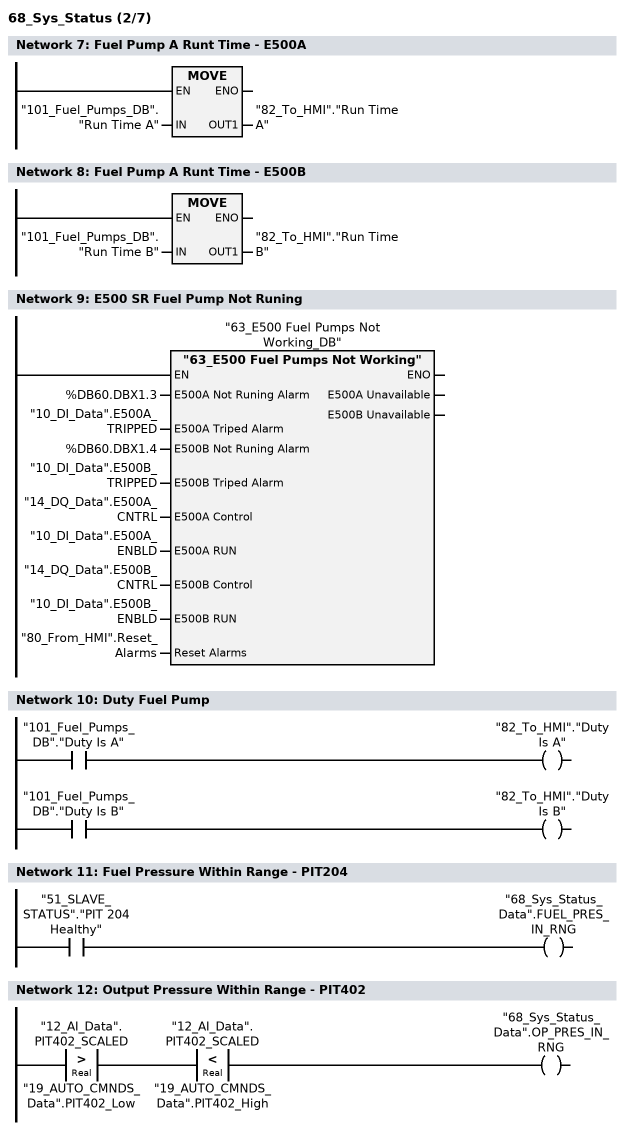
   RUNG wire#powerrail
      Move(in := "101_Fuel_Pumps_DB"."Run Time A", out1 => "82_To_HMI"."Run Time A")
   END_RUNG
   // the same network as SCL:
   "82_To_HMI"."Run Time A" := "101_Fuel_Pumps_DB"."Run Time A";
END_REGION

REGION Network 8: Fuel Pump A Runt Time - E500B
   RUNG wire#powerrail
      Move(in := "101_Fuel_Pumps_DB"."Run Time B", out1 => "82_To_HMI"."Run Time B")
   END_RUNG
   // the same network as SCL:
   "82_To_HMI"."Run Time B" := "101_Fuel_Pumps_DB"."Run Time B";
END_REGION

REGION Network 9: E500 SR Fuel Pump Not Runing
   RUNG wire#powerrail
      "63_E500 Fuel Pumps Not Working_DB"("E500A Not Runing Alarm" := %DB60.DBX1.3, "E500A Triped Alarm" := "10_DI_Data".E500A_TRIPPED, "E500B Not Runing Alarm" := %DB60.DBX1.4, "E500B Triped Alarm" := "10_DI_Data".E500B_TRIPPED, "E500A Control" := "14_DQ_Data".E500A_CNTRL, "E500A RUN" := "10_DI_Data".E500A_ENBLD, "E500B Control" := "14_DQ_Data".E500B_CNTRL, "E500B RUN" := "10_DI_Data".E500B_ENBLD, "Reset Alarms" := "80_From_HMI".Reset_Alarms, "E500A Unavailable" =>, "E500B Unavailable" =>)
   END_RUNG
   // the same network as SCL:
   "63_E500 Fuel Pumps Not Working_DB"("E500A Not Runing Alarm" := %DB60.DBX1.3,   // "63_E500 Fuel Pumps Not Working"
                           "E500A Triped Alarm" := "10_DI_Data".E500A_TRIPPED,
                           "E500B Not Runing Alarm" := %DB60.DBX1.4,
                           "E500B Triped Alarm" := "10_DI_Data".E500B_TRIPPED,
                           "E500A Control" := "14_DQ_Data".E500A_CNTRL,
                           "E500A RUN" := "10_DI_Data".E500A_ENBLD,
                           "E500B Control" := "14_DQ_Data".E500B_CNTRL,
                           "E500B RUN" := "10_DI_Data".E500B_ENBLD,
                           "Reset Alarms" := "80_From_HMI".Reset_Alarms);
END_REGION

REGION Network 10: Duty Fuel Pump
   RUNG wire#powerrail
      Contact( "101_Fuel_Pumps_DB"."Duty Is A" )
      Coil( "82_To_HMI"."Duty Is A" )
   END_RUNG
   RUNG wire#powerrail
      Contact( "101_Fuel_Pumps_DB"."Duty Is B" )
      Coil( "82_To_HMI"."Duty Is B" )
   END_RUNG
   // the same network as SCL:
   "82_To_HMI"."Duty Is A" := "101_Fuel_Pumps_DB"."Duty Is A";
   "82_To_HMI"."Duty Is B" := "101_Fuel_Pumps_DB"."Duty Is B";
END_REGION

REGION Network 11: Fuel Pressure Within Range - PIT204
   RUNG wire#powerrail
      Contact( "51_SLAVE_STATUS"."PIT 204 Healthy" )
      Coil( "68_Sys_Status_Data".FUEL_PRES_IN_RNG )
   END_RUNG
   // the same network as SCL:
   "68_Sys_Status_Data".FUEL_PRES_IN_RNG := "51_SLAVE_STATUS"."PIT 204 Healthy";
END_REGION

REGION Network 12: Output Pressure Within Range - PIT402
   RUNG wire#powerrail
      { S7_Templates := "SrcType := Real" } GT_Contact(in1 := "12_AI_Data".PIT402_SCALED, in2 := "19_AUTO_CMNDS_Data".PIT402_Low)
      { S7_Templates := "SrcType := Real" } LT_Contact(in1 := "12_AI_Data".PIT402_SCALED, in2 := "19_AUTO_CMNDS_Data".PIT402_High)
      Coil( "68_Sys_Status_Data".OP_PRES_IN_RNG )
   END_RUNG
   // the same network as SCL:
   "68_Sys_Status_Data".OP_PRES_IN_RNG := ("12_AI_Data".PIT402_SCALED > "19_AUTO_CMNDS_Data".PIT402_Low) AND ("12_AI_Data".PIT402_SCALED < "19_AUTO_CMNDS_Data".PIT402_High);
END_REGION

REGION Network 13: Cargo Banketing Mode
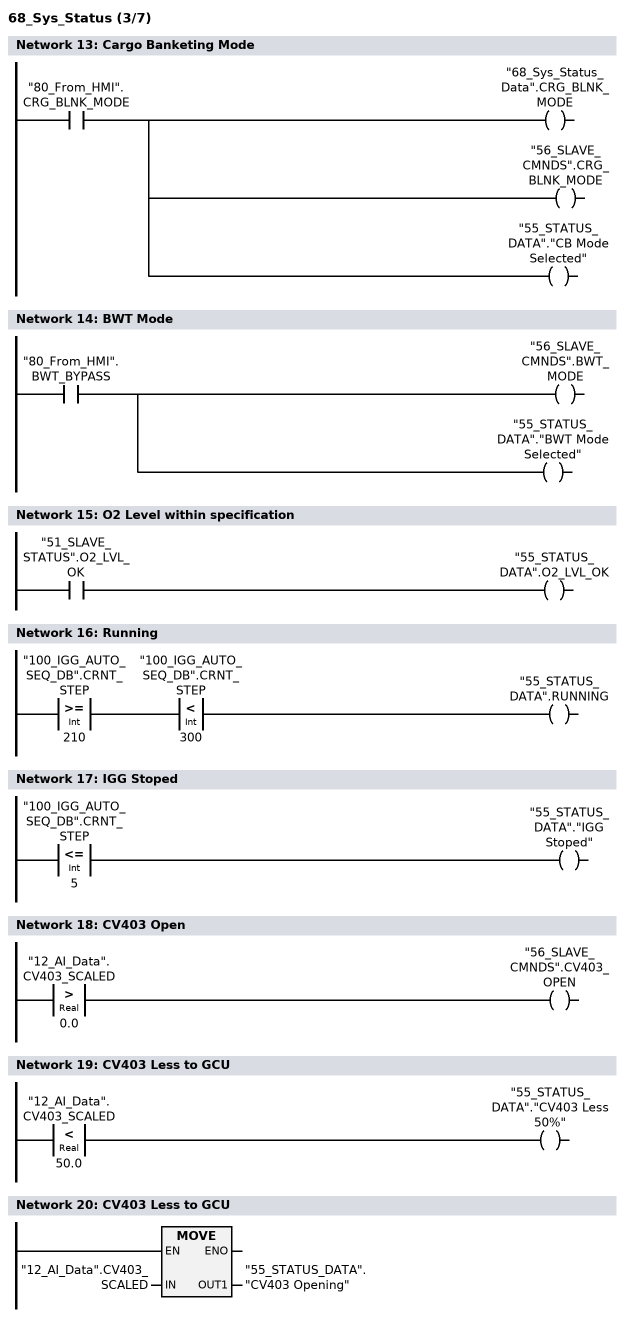
   RUNG wire#powerrail
      Contact( "80_From_HMI".CRG_BLNK_MODE )
      wire#w1
      Coil( "68_Sys_Status_Data".CRG_BLNK_MODE )
   END_RUNG
   RUNG wire#w1
      Coil( "56_SLAVE_CMNDS".CRG_BLNK_MODE )
   END_RUNG
   RUNG wire#w1
      Coil( "55_STATUS_DATA"."CB Mode Selected" )
   END_RUNG
   // the same network as SCL:
   "68_Sys_Status_Data".CRG_BLNK_MODE := "80_From_HMI".CRG_BLNK_MODE;
   "56_SLAVE_CMNDS".CRG_BLNK_MODE := "80_From_HMI".CRG_BLNK_MODE;
   "55_STATUS_DATA"."CB Mode Selected" := "80_From_HMI".CRG_BLNK_MODE;
END_REGION

REGION Network 14: BWT Mode
   RUNG wire#powerrail
      Contact( "80_From_HMI".BWT_BYPASS )
      wire#w1
      Coil( "56_SLAVE_CMNDS".BWT_MODE )
   END_RUNG
   RUNG wire#w1
      Coil( "55_STATUS_DATA"."BWT Mode Selected" )
   END_RUNG
   // the same network as SCL:
   "56_SLAVE_CMNDS".BWT_MODE := "80_From_HMI".BWT_BYPASS;
   "55_STATUS_DATA"."BWT Mode Selected" := "80_From_HMI".BWT_BYPASS;
END_REGION

REGION Network 15: O2 Level within specification
   RUNG wire#powerrail
      Contact( "51_SLAVE_STATUS".O2_LVL_OK )
      Coil( "55_STATUS_DATA".O2_LVL_OK )
   END_RUNG
   // the same network as SCL:
   "55_STATUS_DATA".O2_LVL_OK := "51_SLAVE_STATUS".O2_LVL_OK;
END_REGION

REGION Network 16: Running
   RUNG wire#powerrail
      { S7_Templates := "SrcType := Int" } GE_Contact(in1 := "100_IGG_AUTO_SEQ_DB".CRNT_STEP, in2 := 210)
      { S7_Templates := "SrcType := Int" } LT_Contact(in1 := "100_IGG_AUTO_SEQ_DB".CRNT_STEP, in2 := 300)
      Coil( "55_STATUS_DATA".RUNNING )
   END_RUNG
   // the same network as SCL:
   "55_STATUS_DATA".RUNNING := ("100_IGG_AUTO_SEQ_DB".CRNT_STEP >= 210) AND ("100_IGG_AUTO_SEQ_DB".CRNT_STEP < 300);
END_REGION

REGION Network 17: IGG Stoped
   RUNG wire#powerrail
      { S7_Templates := "SrcType := Int" } LE_Contact(in1 := "100_IGG_AUTO_SEQ_DB".CRNT_STEP, in2 := 5)
      Coil( "55_STATUS_DATA"."IGG Stoped" )
   END_RUNG
   // the same network as SCL:
   "55_STATUS_DATA"."IGG Stoped" := "100_IGG_AUTO_SEQ_DB".CRNT_STEP <= 5;
END_REGION

REGION Network 18: CV403 Open
   RUNG wire#powerrail
      { S7_Templates := "SrcType := Real" } GT_Contact(in1 := "12_AI_Data".CV403_SCALED, in2 := 0.0)
      Coil( "56_SLAVE_CMNDS".CV403_OPEN )
   END_RUNG
   // the same network as SCL:
   "56_SLAVE_CMNDS".CV403_OPEN := "12_AI_Data".CV403_SCALED > 0.0;
END_REGION

REGION Network 19: CV403 Less to GCU
   RUNG wire#powerrail
      { S7_Templates := "SrcType := Real" } LT_Contact(in1 := "12_AI_Data".CV403_SCALED, in2 := 50.0)
      Coil( "55_STATUS_DATA"."CV403 Less 50%" )
   END_RUNG
   // the same network as SCL:
   "55_STATUS_DATA"."CV403 Less 50%" := "12_AI_Data".CV403_SCALED < 50.0;
END_REGION

REGION Network 20: CV403 Less to GCU
   RUNG wire#powerrail
      Move(in := "12_AI_Data".CV403_SCALED, out1 => "55_STATUS_DATA"."CV403 Opening")
   END_RUNG
   // the same network as SCL:
   "55_STATUS_DATA"."CV403 Opening" := "12_AI_Data".CV403_SCALED;
END_REGION

REGION Network 21: Fuel Pump 1 Enabled E500A
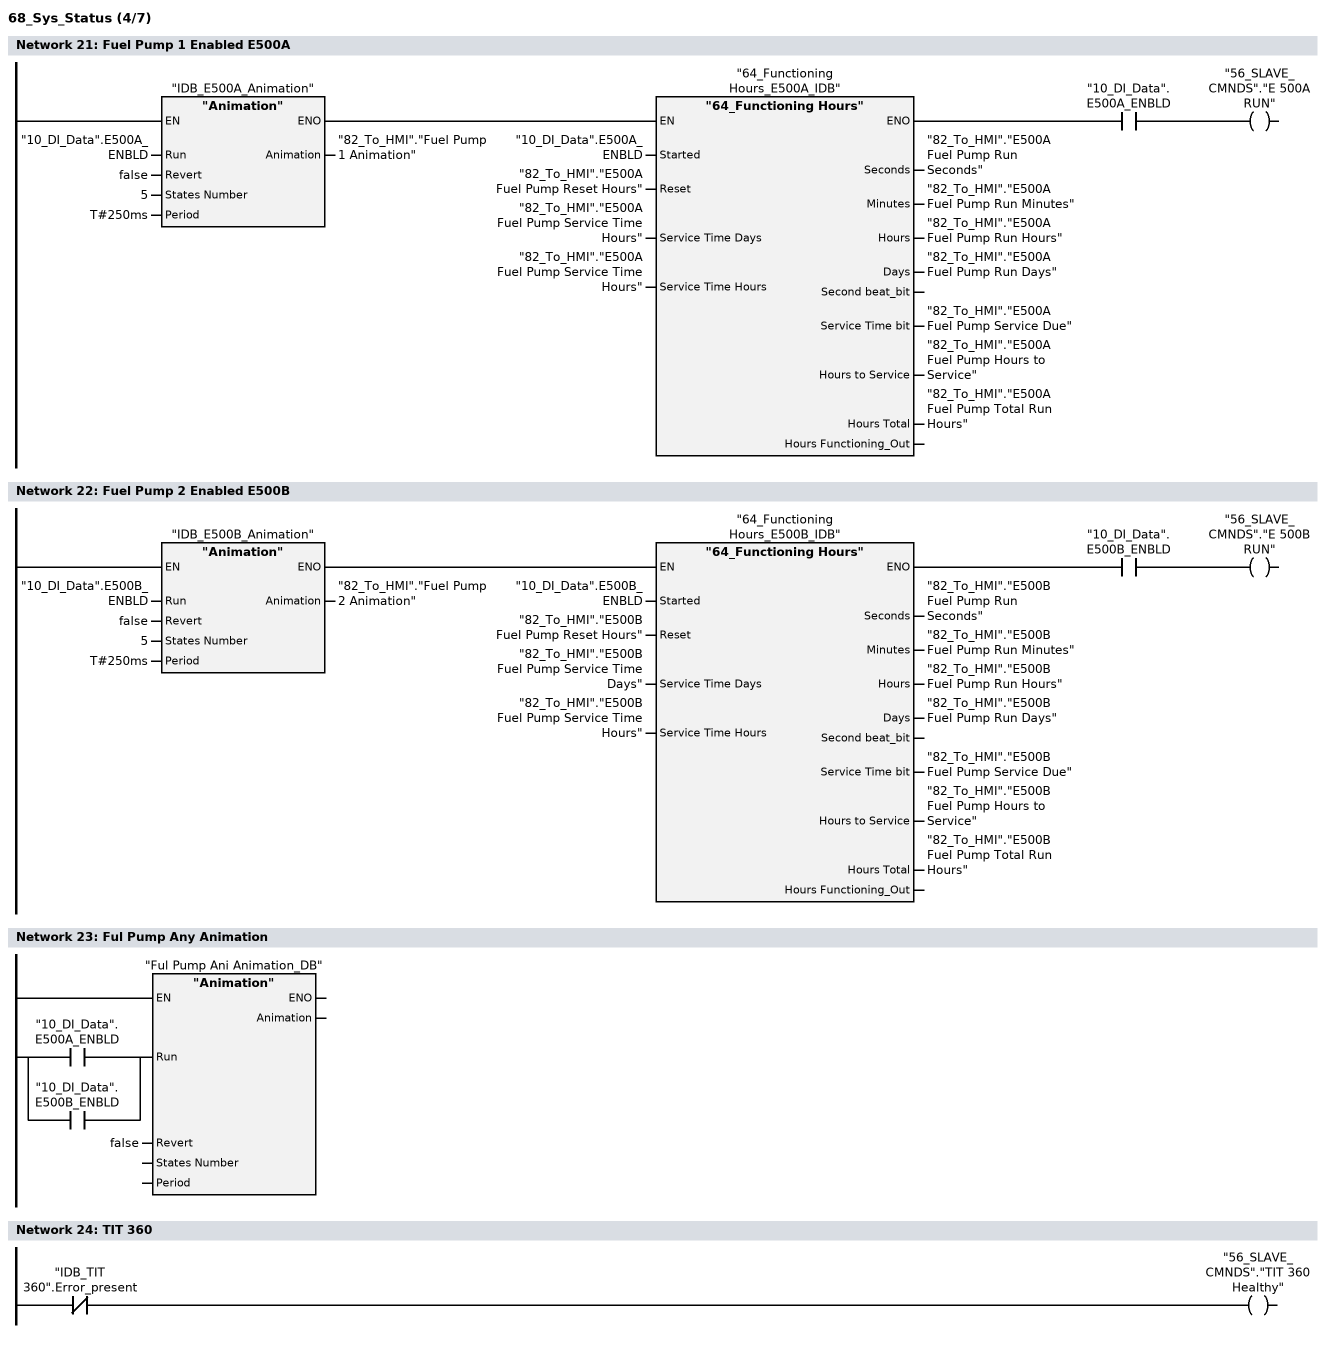
   RUNG wire#powerrail
      "IDB_E500A_Animation"(Run := "10_DI_Data".E500A_ENBLD, Revert := false, "States Number" := 5, Period := T#250ms, Animation => "82_To_HMI"."Fuel Pump 1 Animation")
      "64_Functioning Hours_E500A_IDB"(Started := "10_DI_Data".E500A_ENBLD, Reset := "82_To_HMI"."E500A Fuel Pump Reset Hours", "Service Time Days" := "82_To_HMI"."E500A Fuel Pump Service Time Hours", "Service Time Hours" := "82_To_HMI"."E500A Fuel Pump Service Time Hours", Seconds => "82_To_HMI"."E500A Fuel Pump Run Seconds", Minutes => "82_To_HMI"."E500A Fuel Pump Run Minutes", Hours => "82_To_HMI"."E500A Fuel Pump Run Hours", Days => "82_To_HMI"."E500A Fuel Pump Run Days", "Second beat_bit" =>, "Service Time bit" => "82_To_HMI"."E500A Fuel Pump Service Due", "Hours to Service" => "82_To_HMI"."E500A Fuel Pump Hours to Service", "Hours Total" => "82_To_HMI"."E500A Fuel Pump Total Run Hours", "Hours Functioning_Out" =>)
      Contact( "10_DI_Data".E500A_ENBLD )
      Coil( "56_SLAVE_CMNDS"."E 500A RUN" )
   END_RUNG
   // the same network as SCL:
   "IDB_E500A_Animation"(Run := "10_DI_Data".E500A_ENBLD,   // "Animation"
                         Revert := false,
                         "States Number" := 5,
                         Period := T#250ms,
                         Animation => "82_To_HMI"."Fuel Pump 1 Animation",
                         ENO => #_w1);
   "64_Functioning Hours_E500A_IDB"(EN := #_w1,   // "64_Functioning Hours"
                           Started := "10_DI_Data".E500A_ENBLD,
                           Reset := "82_To_HMI"."E500A Fuel Pump Reset Hours",
                           "Service Time Days" := "82_To_HMI"."E500A Fuel Pump Service Time Hours",
                           "Service Time Hours" := "82_To_HMI"."E500A Fuel Pump Service Time Hours",
                           Seconds => "82_To_HMI"."E500A Fuel Pump Run Seconds",
                           Minutes => "82_To_HMI"."E500A Fuel Pump Run Minutes",
                           Hours => "82_To_HMI"."E500A Fuel Pump Run Hours",
                           Days => "82_To_HMI"."E500A Fuel Pump Run Days",
                           "Service Time bit" => "82_To_HMI"."E500A Fuel Pump Service Due",
                           "Hours to Service" => "82_To_HMI"."E500A Fuel Pump Hours to Service",
                           "Hours Total" => "82_To_HMI"."E500A Fuel Pump Total Run Hours",
                           ENO => #_w2);
   "56_SLAVE_CMNDS"."E 500A RUN" := #_w2 AND "10_DI_Data".E500A_ENBLD;
END_REGION

REGION Network 22: Fuel Pump 2 Enabled E500B
   RUNG wire#powerrail
      "IDB_E500B_Animation"(Run := "10_DI_Data".E500B_ENBLD, Revert := false, "States Number" := 5, Period := T#250ms, Animation => "82_To_HMI"."Fuel Pump 2 Animation")
      "64_Functioning Hours_E500B_IDB"(Started := "10_DI_Data".E500B_ENBLD, Reset := "82_To_HMI"."E500B Fuel Pump Reset Hours", "Service Time Days" := "82_To_HMI"."E500B Fuel Pump Service Time Days", "Service Time Hours" := "82_To_HMI"."E500B Fuel Pump Service Time Hours", Seconds => "82_To_HMI"."E500B Fuel Pump Run Seconds", Minutes => "82_To_HMI"."E500B Fuel Pump Run Minutes", Hours => "82_To_HMI"."E500B Fuel Pump Run Hours", Days => "82_To_HMI"."E500B Fuel Pump Run Days", "Second beat_bit" =>, "Service Time bit" => "82_To_HMI"."E500B Fuel Pump Service Due", "Hours to Service" => "82_To_HMI"."E500B Fuel Pump Hours to Service", "Hours Total" => "82_To_HMI"."E500B Fuel Pump Total Run Hours", "Hours Functioning_Out" =>)
      Contact( "10_DI_Data".E500B_ENBLD )
      Coil( "56_SLAVE_CMNDS"."E 500B RUN" )
   END_RUNG
   // the same network as SCL:
   "IDB_E500B_Animation"(Run := "10_DI_Data".E500B_ENBLD,   // "Animation"
                         Revert := false,
                         "States Number" := 5,
                         Period := T#250ms,
                         Animation => "82_To_HMI"."Fuel Pump 2 Animation",
                         ENO => #_w1);
   "64_Functioning Hours_E500B_IDB"(EN := #_w1,   // "64_Functioning Hours"
                           Started := "10_DI_Data".E500B_ENBLD,
                           Reset := "82_To_HMI"."E500B Fuel Pump Reset Hours",
                           "Service Time Days" := "82_To_HMI"."E500B Fuel Pump Service Time Days",
                           "Service Time Hours" := "82_To_HMI"."E500B Fuel Pump Service Time Hours",
                           Seconds => "82_To_HMI"."E500B Fuel Pump Run Seconds",
                           Minutes => "82_To_HMI"."E500B Fuel Pump Run Minutes",
                           Hours => "82_To_HMI"."E500B Fuel Pump Run Hours",
                           Days => "82_To_HMI"."E500B Fuel Pump Run Days",
                           "Service Time bit" => "82_To_HMI"."E500B Fuel Pump Service Due",
                           "Hours to Service" => "82_To_HMI"."E500B Fuel Pump Hours to Service",
                           "Hours Total" => "82_To_HMI"."E500B Fuel Pump Total Run Hours",
                           ENO => #_w2);
   "56_SLAVE_CMNDS"."E 500B RUN" := #_w2 AND "10_DI_Data".E500B_ENBLD;
END_REGION

REGION Network 23: Ful Pump Any Animation
   RUNG wire#powerrail
      "Ful Pump Ani Animation_DB"(Run := wire#w1, Revert := false, "States Number" :=, Period :=, Animation =>)
   END_RUNG
   RUNG wire#powerrail
      Contact( "10_DI_Data".E500A_ENBLD )
   END_RUNG wire#w1
   RUNG wire#powerrail
      Contact( "10_DI_Data".E500B_ENBLD )
   END_RUNG wire#w1
   // the same network as SCL:
   "Ful Pump Ani Animation_DB"(Run := "10_DI_Data".E500A_ENBLD OR "10_DI_Data".E500B_ENBLD, Revert := false);   // "Animation"
END_REGION

REGION Network 24: TIT 360
   RUNG wire#powerrail
      I_Contact( "IDB_TIT 360".Error_present )
      Coil( "56_SLAVE_CMNDS"."TIT 360 Healthy" )
   END_RUNG
   // the same network as SCL:
   "56_SLAVE_CMNDS"."TIT 360 Healthy" := NOT "IDB_TIT 360".Error_present;
END_REGION

REGION Network 25: TIT 401
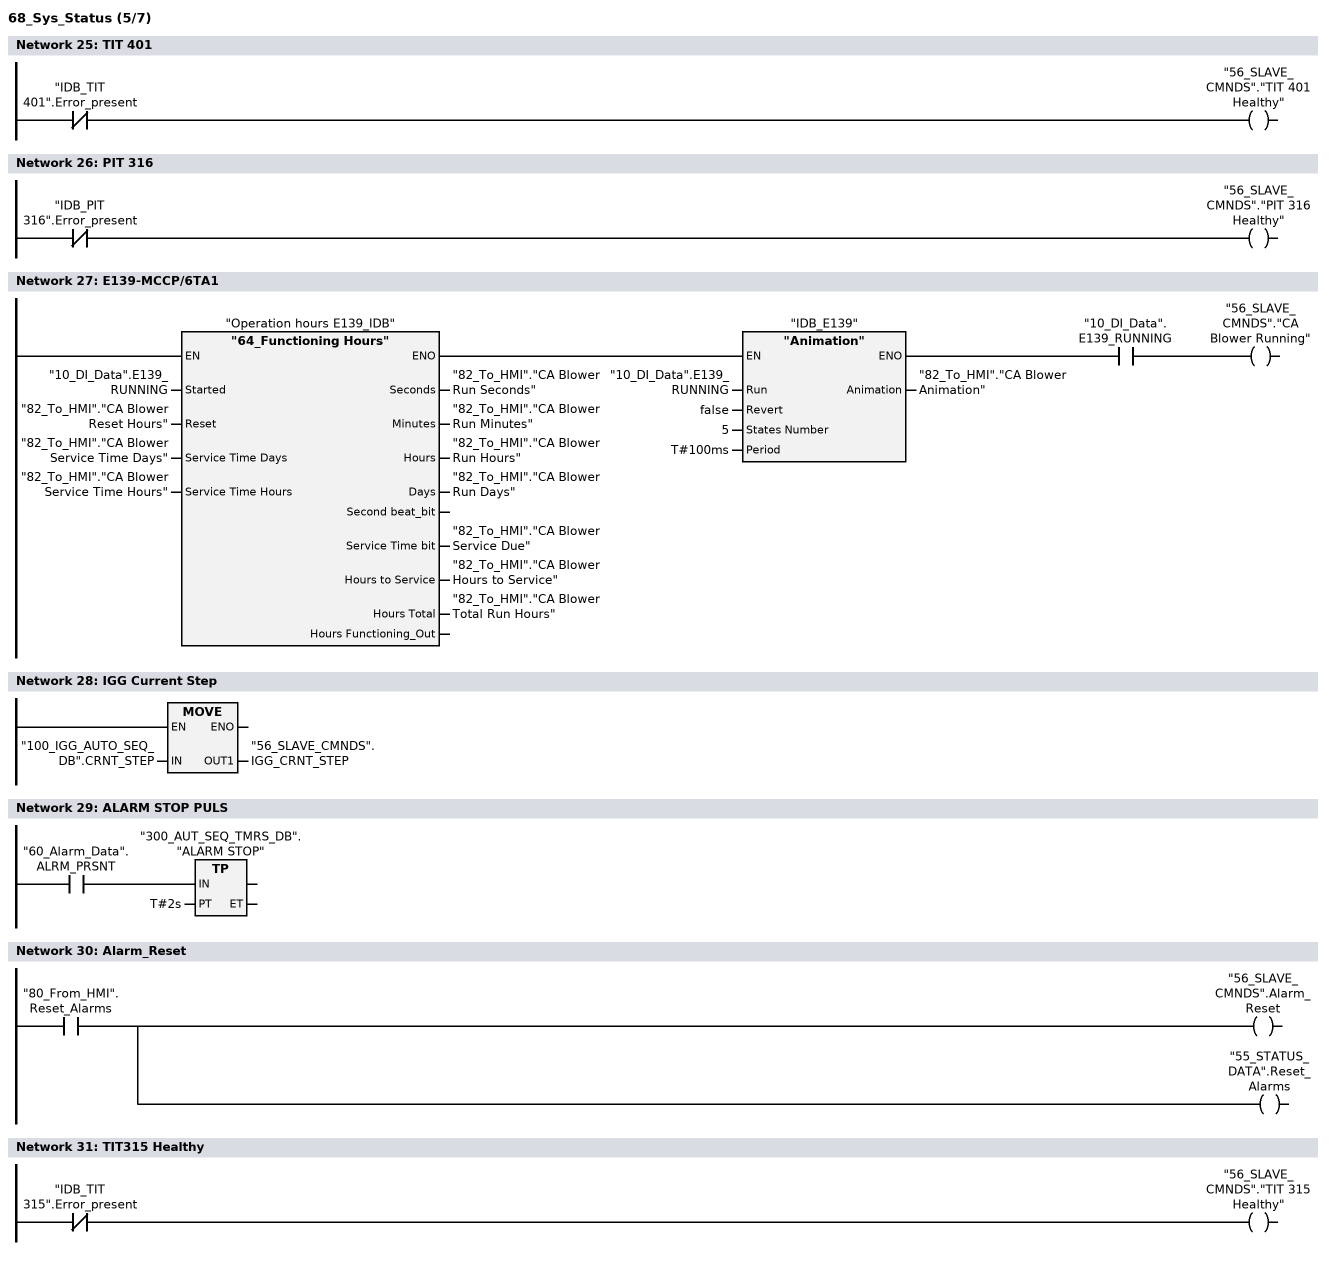
   RUNG wire#powerrail
      I_Contact( "IDB_TIT 401".Error_present )
      Coil( "56_SLAVE_CMNDS"."TIT 401 Healthy" )
   END_RUNG
   // the same network as SCL:
   "56_SLAVE_CMNDS"."TIT 401 Healthy" := NOT "IDB_TIT 401".Error_present;
END_REGION

REGION Network 26: PIT 316
   RUNG wire#powerrail
      I_Contact( "IDB_PIT 316".Error_present )
      Coil( "56_SLAVE_CMNDS"."PIT 316 Healthy" )
   END_RUNG
   // the same network as SCL:
   "56_SLAVE_CMNDS"."PIT 316 Healthy" := NOT "IDB_PIT 316".Error_present;
END_REGION

REGION Network 27: E139-MCCP/6TA1
   RUNG wire#powerrail
      "Operation hours E139_IDB"(Started := "10_DI_Data".E139_RUNNING, Reset := "82_To_HMI"."CA Blower Reset Hours", "Service Time Days" := "82_To_HMI"."CA Blower Service Time Days", "Service Time Hours" := "82_To_HMI"."CA Blower Service Time Hours", Seconds => "82_To_HMI"."CA Blower Run Seconds", Minutes => "82_To_HMI"."CA Blower Run Minutes", Hours => "82_To_HMI"."CA Blower Run Hours", Days => "82_To_HMI"."CA Blower Run Days", "Second beat_bit" =>, "Service Time bit" => "82_To_HMI"."CA Blower Service Due", "Hours to Service" => "82_To_HMI"."CA Blower Hours to Service", "Hours Total" => "82_To_HMI"."CA Blower Total Run Hours", "Hours Functioning_Out" =>)
      "IDB_E139"(Run := "10_DI_Data".E139_RUNNING, Revert := false, "States Number" := 5, Period := T#100ms, Animation => "82_To_HMI"."CA Blower Animation")
      Contact( "10_DI_Data".E139_RUNNING )
      Coil( "56_SLAVE_CMNDS"."CA Blower Running" )
   END_RUNG
   // the same network as SCL:
   "Operation hours E139_IDB"(Started := "10_DI_Data".E139_RUNNING,   // "64_Functioning Hours"
                           Reset := "82_To_HMI"."CA Blower Reset Hours",
                           "Service Time Days" := "82_To_HMI"."CA Blower Service Time Days",
                           "Service Time Hours" := "82_To_HMI"."CA Blower Service Time Hours",
                           Seconds => "82_To_HMI"."CA Blower Run Seconds",
                           Minutes => "82_To_HMI"."CA Blower Run Minutes",
                           Hours => "82_To_HMI"."CA Blower Run Hours",
                           Days => "82_To_HMI"."CA Blower Run Days",
                           "Service Time bit" => "82_To_HMI"."CA Blower Service Due",
                           "Hours to Service" => "82_To_HMI"."CA Blower Hours to Service",
                           "Hours Total" => "82_To_HMI"."CA Blower Total Run Hours",
                           ENO => #_w1);
   "IDB_E139"(EN := #_w1,   // "Animation"
              Run := "10_DI_Data".E139_RUNNING,
              Revert := false,
              "States Number" := 5,
              Period := T#100ms,
              Animation => "82_To_HMI"."CA Blower Animation",
              ENO => #_w2);
   "56_SLAVE_CMNDS"."CA Blower Running" := #_w2 AND "10_DI_Data".E139_RUNNING;
END_REGION

REGION Network 28: IGG Current Step
   RUNG wire#powerrail
      Move(in := "100_IGG_AUTO_SEQ_DB".CRNT_STEP, out1 => "56_SLAVE_CMNDS".IGG_CRNT_STEP)
   END_RUNG
   // the same network as SCL:
   "56_SLAVE_CMNDS".IGG_CRNT_STEP := "100_IGG_AUTO_SEQ_DB".CRNT_STEP;
END_REGION

REGION Network 29: ALARM STOP PULS
   "300_AUT_SEQ_TMRS_DB"."ALARM STOP".TP(IN := "60_Alarm_Data".ALRM_PRSNT, PT := T#2s);
END_REGION

REGION Network 30: Alarm_Reset
   RUNG wire#powerrail
      Contact( "80_From_HMI".Reset_Alarms )
      wire#w1
      Coil( "56_SLAVE_CMNDS".Alarm_Reset )
   END_RUNG
   RUNG wire#w1
      Coil( "55_STATUS_DATA".Reset_Alarms )
   END_RUNG
   // the same network as SCL:
   "56_SLAVE_CMNDS".Alarm_Reset := "80_From_HMI".Reset_Alarms;
   "55_STATUS_DATA".Reset_Alarms := "80_From_HMI".Reset_Alarms;
END_REGION

REGION Network 31: TIT315 Healthy
   RUNG wire#powerrail
      I_Contact( "IDB_TIT 315".Error_present )
      Coil( "56_SLAVE_CMNDS"."TIT 315 Healthy" )
   END_RUNG
   // the same network as SCL:
   "56_SLAVE_CMNDS"."TIT 315 Healthy" := NOT "IDB_TIT 315".Error_present;
END_REGION

REGION Network 32: Safety System Interlock SFTY_SYS_IL
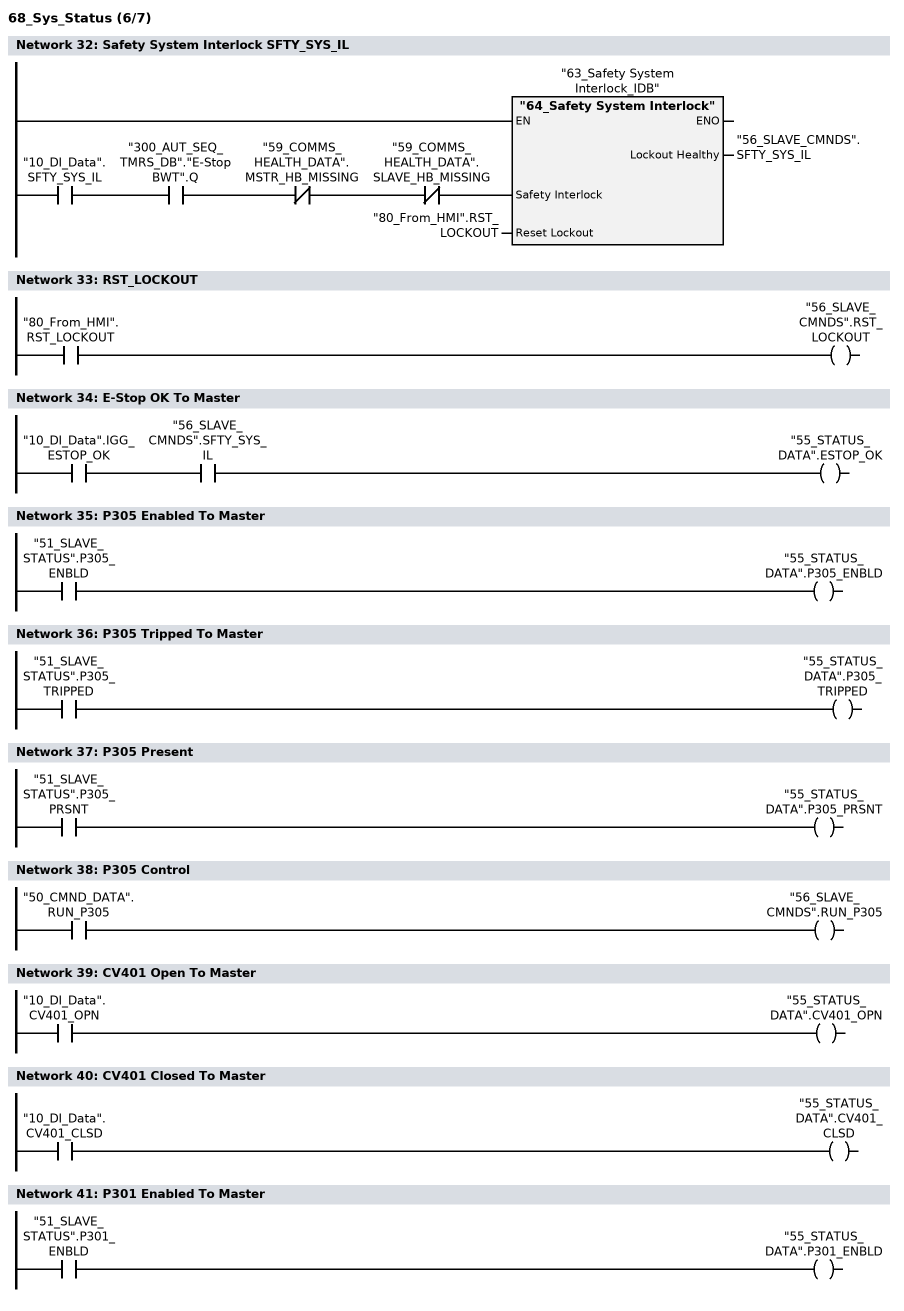
   RUNG wire#powerrail
      "63_Safety System Interlock_IDB"("Safety Interlock" := wire#w1, "Reset Lockout" := "80_From_HMI".RST_LOCKOUT, "Lockout Healthy" => "56_SLAVE_CMNDS".SFTY_SYS_IL)
   END_RUNG
   RUNG wire#powerrail
      Contact( "10_DI_Data".SFTY_SYS_IL )
      Contact( "300_AUT_SEQ_TMRS_DB"."E-Stop BWT".Q )
      I_Contact( "59_COMMS_HEALTH_DATA".MSTR_HB_MISSING )
      I_Contact( "59_COMMS_HEALTH_DATA".SLAVE_HB_MISSING )
   END_RUNG wire#w1
   // the same network as SCL:
   "63_Safety System Interlock_IDB"("Safety Interlock" := "10_DI_Data".SFTY_SYS_IL AND "300_AUT_SEQ_TMRS_DB"."E-Stop BWT".Q AND NOT "59_COMMS_HEALTH_DATA".MSTR_HB_MISSING AND NOT "59_COMMS_HEALTH_DATA".SLAVE_HB_MISSING,   // "64_Safety System Interlock"
                           "Reset Lockout" := "80_From_HMI".RST_LOCKOUT,
                           "Lockout Healthy" => "56_SLAVE_CMNDS".SFTY_SYS_IL);
END_REGION

REGION Network 33: RST_LOCKOUT
   RUNG wire#powerrail
      Contact( "80_From_HMI".RST_LOCKOUT )
      Coil( "56_SLAVE_CMNDS".RST_LOCKOUT )
   END_RUNG
   // the same network as SCL:
   "56_SLAVE_CMNDS".RST_LOCKOUT := "80_From_HMI".RST_LOCKOUT;
END_REGION

REGION Network 34: E-Stop OK To Master
   RUNG wire#powerrail
      Contact( "10_DI_Data".IGG_ESTOP_OK )
      Contact( "56_SLAVE_CMNDS".SFTY_SYS_IL )
      Coil( "55_STATUS_DATA".ESTOP_OK )
   END_RUNG
   // the same network as SCL:
   "55_STATUS_DATA".ESTOP_OK := "10_DI_Data".IGG_ESTOP_OK AND "56_SLAVE_CMNDS".SFTY_SYS_IL;
END_REGION

REGION Network 35: P305 Enabled To Master
   RUNG wire#powerrail
      Contact( "51_SLAVE_STATUS".P305_ENBLD )
      Coil( "55_STATUS_DATA".P305_ENBLD )
   END_RUNG
   // the same network as SCL:
   "55_STATUS_DATA".P305_ENBLD := "51_SLAVE_STATUS".P305_ENBLD;
END_REGION

REGION Network 36: P305 Tripped To Master
   RUNG wire#powerrail
      Contact( "51_SLAVE_STATUS".P305_TRIPPED )
      Coil( "55_STATUS_DATA".P305_TRIPPED )
   END_RUNG
   // the same network as SCL:
   "55_STATUS_DATA".P305_TRIPPED := "51_SLAVE_STATUS".P305_TRIPPED;
END_REGION

REGION Network 37: P305 Present
   RUNG wire#powerrail
      Contact( "51_SLAVE_STATUS".P305_PRSNT )
      Coil( "55_STATUS_DATA".P305_PRSNT )
   END_RUNG
   // the same network as SCL:
   "55_STATUS_DATA".P305_PRSNT := "51_SLAVE_STATUS".P305_PRSNT;
END_REGION

REGION Network 38: P305 Control
   RUNG wire#powerrail
      Contact( "50_CMND_DATA".RUN_P305 )
      Coil( "56_SLAVE_CMNDS".RUN_P305 )
   END_RUNG
   // the same network as SCL:
   "56_SLAVE_CMNDS".RUN_P305 := "50_CMND_DATA".RUN_P305;
END_REGION

REGION Network 39: CV401 Open To Master
   RUNG wire#powerrail
      Contact( "10_DI_Data".CV401_OPN )
      Coil( "55_STATUS_DATA".CV401_OPN )
   END_RUNG
   // the same network as SCL:
   "55_STATUS_DATA".CV401_OPN := "10_DI_Data".CV401_OPN;
END_REGION

REGION Network 40: CV401 Closed To Master
   RUNG wire#powerrail
      Contact( "10_DI_Data".CV401_CLSD )
      Coil( "55_STATUS_DATA".CV401_CLSD )
   END_RUNG
   // the same network as SCL:
   "55_STATUS_DATA".CV401_CLSD := "10_DI_Data".CV401_CLSD;
END_REGION

REGION Network 41: P301 Enabled To Master
   RUNG wire#powerrail
      Contact( "51_SLAVE_STATUS".P301_ENBLD )
      Coil( "55_STATUS_DATA".P301_ENBLD )
   END_RUNG
   // the same network as SCL:
   "55_STATUS_DATA".P301_ENBLD := "51_SLAVE_STATUS".P301_ENBLD;
END_REGION

REGION Network 42: CV311 Open To Master
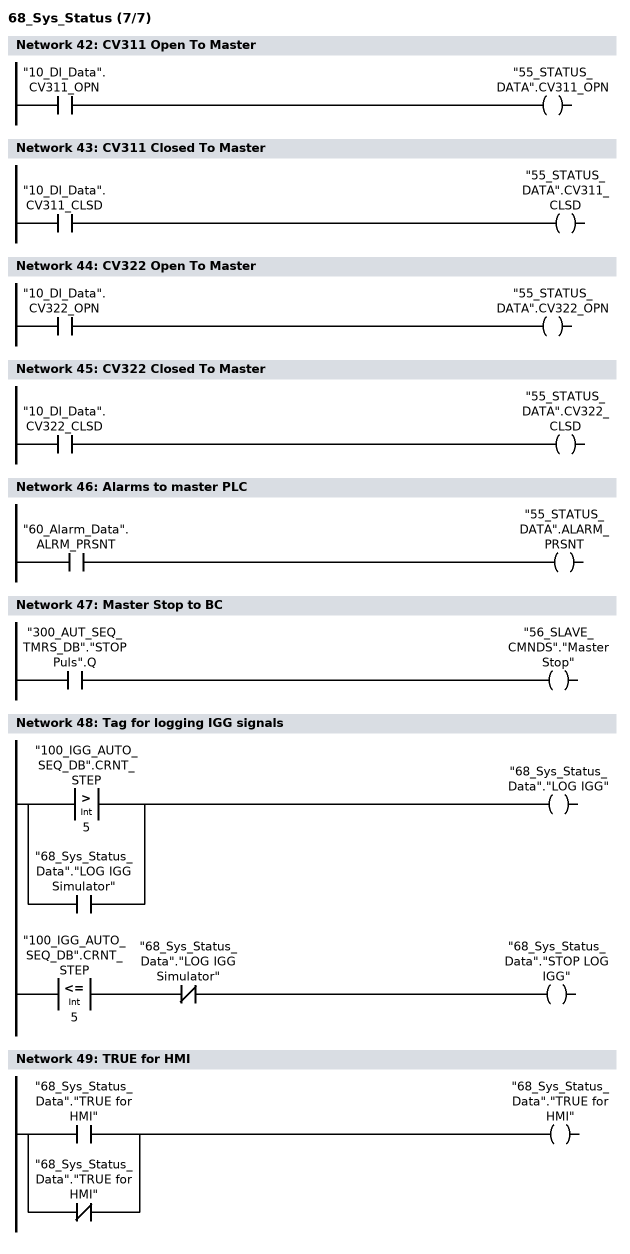
   RUNG wire#powerrail
      Contact( "10_DI_Data".CV311_OPN )
      Coil( "55_STATUS_DATA".CV311_OPN )
   END_RUNG
   // the same network as SCL:
   "55_STATUS_DATA".CV311_OPN := "10_DI_Data".CV311_OPN;
END_REGION

REGION Network 43: CV311 Closed To Master
   RUNG wire#powerrail
      Contact( "10_DI_Data".CV311_CLSD )
      Coil( "55_STATUS_DATA".CV311_CLSD )
   END_RUNG
   // the same network as SCL:
   "55_STATUS_DATA".CV311_CLSD := "10_DI_Data".CV311_CLSD;
END_REGION

REGION Network 44: CV322 Open To Master
   RUNG wire#powerrail
      Contact( "10_DI_Data".CV322_OPN )
      Coil( "55_STATUS_DATA".CV322_OPN )
   END_RUNG
   // the same network as SCL:
   "55_STATUS_DATA".CV322_OPN := "10_DI_Data".CV322_OPN;
END_REGION

REGION Network 45: CV322 Closed To Master
   RUNG wire#powerrail
      Contact( "10_DI_Data".CV322_CLSD )
      Coil( "55_STATUS_DATA".CV322_CLSD )
   END_RUNG
   // the same network as SCL:
   "55_STATUS_DATA".CV322_CLSD := "10_DI_Data".CV322_CLSD;
END_REGION

REGION Network 46: Alarms to master PLC
   RUNG wire#powerrail
      Contact( "60_Alarm_Data".ALRM_PRSNT )
      Coil( "55_STATUS_DATA".ALARM_PRSNT )
   END_RUNG
   // the same network as SCL:
   "55_STATUS_DATA".ALARM_PRSNT := "60_Alarm_Data".ALRM_PRSNT;
END_REGION

REGION Network 47: Master Stop to BC
   RUNG wire#powerrail
      Contact( "300_AUT_SEQ_TMRS_DB"."STOP Puls".Q )
      Coil( "56_SLAVE_CMNDS"."Master Stop" )
   END_RUNG
   // the same network as SCL:
   "56_SLAVE_CMNDS"."Master Stop" := "300_AUT_SEQ_TMRS_DB"."STOP Puls".Q;
END_REGION

REGION Network 48: Tag for logging IGG signals
   RUNG wire#powerrail
      { S7_Templates := "SrcType := Int" } GT_Contact(in1 := "100_IGG_AUTO_SEQ_DB".CRNT_STEP, in2 := 5)
      wire#w1
      Coil( "68_Sys_Status_Data"."LOG IGG" )
   END_RUNG
   RUNG wire#powerrail
      Contact( "68_Sys_Status_Data"."LOG IGG Simulator" )
   END_RUNG wire#w1
   RUNG wire#powerrail
      { S7_Templates := "SrcType := Int" } LE_Contact(in1 := "100_IGG_AUTO_SEQ_DB".CRNT_STEP, in2 := 5)
      I_Contact( "68_Sys_Status_Data"."LOG IGG Simulator" )
      Coil( "68_Sys_Status_Data"."STOP LOG IGG" )
   END_RUNG
   // the same network as SCL:
   "68_Sys_Status_Data"."LOG IGG" := ("100_IGG_AUTO_SEQ_DB".CRNT_STEP > 5) OR "68_Sys_Status_Data"."LOG IGG Simulator";
   "68_Sys_Status_Data"."STOP LOG IGG" := ("100_IGG_AUTO_SEQ_DB".CRNT_STEP <= 5) AND NOT "68_Sys_Status_Data"."LOG IGG Simulator";
END_REGION

REGION Network 49: TRUE for HMI
   RUNG wire#powerrail
      Contact( "68_Sys_Status_Data"."TRUE for HMI" )
      wire#w1
      Coil( "68_Sys_Status_Data"."TRUE for HMI" )
   END_RUNG
   RUNG wire#powerrail
      I_Contact( "68_Sys_Status_Data"."TRUE for HMI" )
   END_RUNG wire#w1
   // the same network as SCL:
   "68_Sys_Status_Data"."TRUE for HMI" := "68_Sys_Status_Data"."TRUE for HMI" OR NOT "68_Sys_Status_Data"."TRUE for HMI";
END_REGION
END_FUNCTION

// folder: 70 - 79 Modes of Operation

FUNCTION "70_Mode_Control" : Void   // FC70, LAD
TITLE = Mode Control
{ S7_Optimized_Access := 'TRUE' }
AUTHOR : JRS
VERSION : 0.1
// To determine the current mode of operation 1=Auto(default), 2=Manual, 3=FatAuto, 4=FatManual
   VAR_TEMP   // added for the SCL form of the ladder/FBD networks
      _w1 : Bool;
   END_VAR
BEGIN

REGION Network 1: Default = Automatic
   // Set default to Automatic (on first scan)
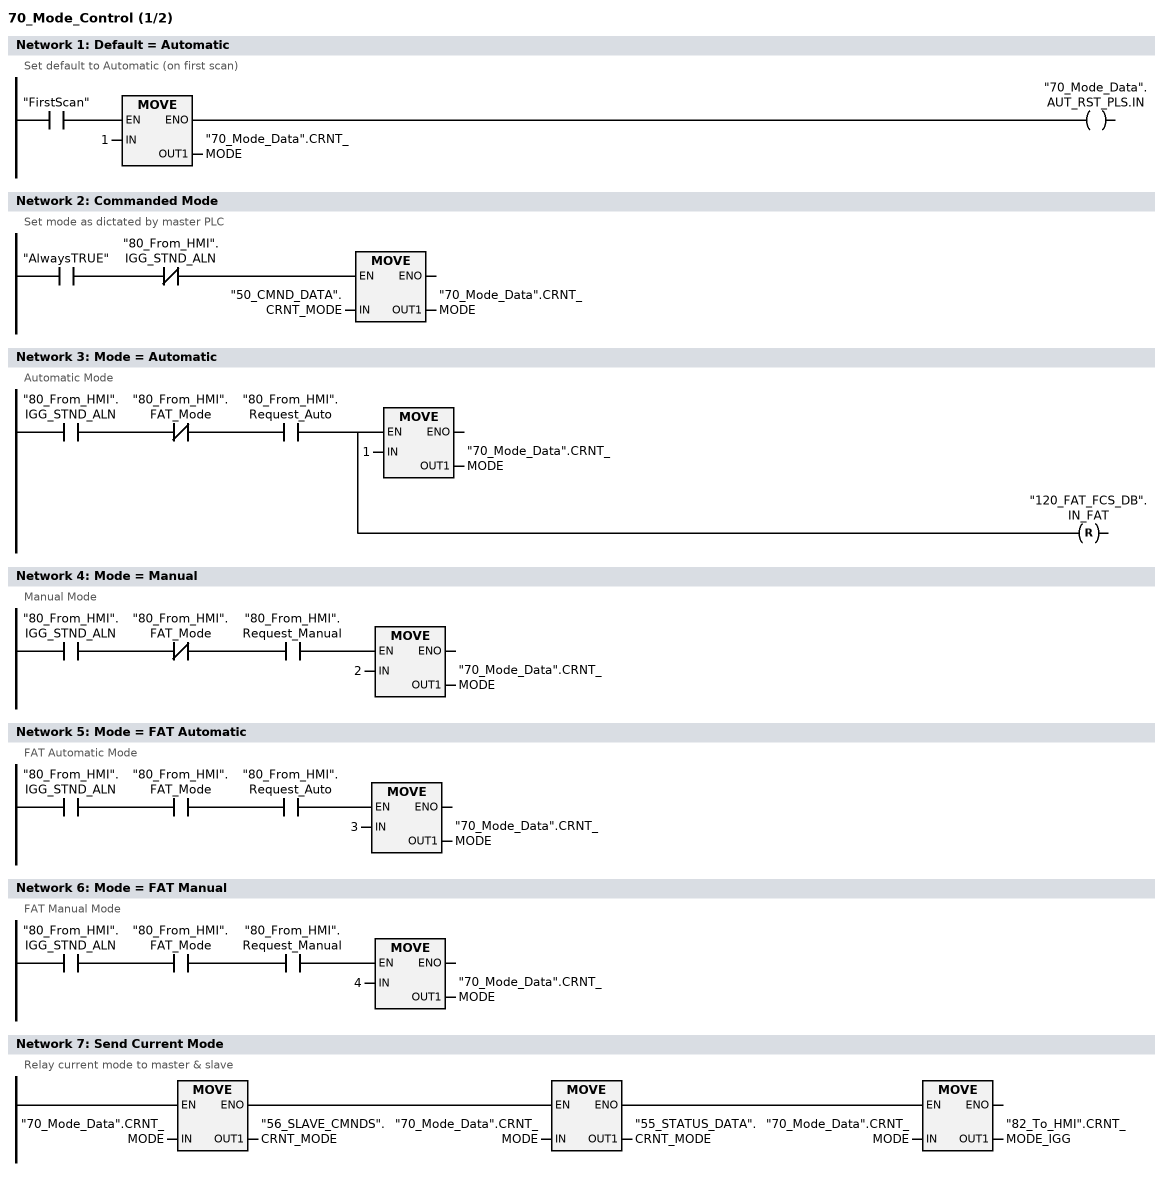
   RUNG wire#powerrail
      Contact( "FirstScan" )
      Move(in := 1, out1 => "70_Mode_Data".CRNT_MODE)
      Coil( "70_Mode_Data".AUT_RST_PLS.IN )
   END_RUNG
   // the same network as SCL:
   IF "FirstScan" THEN "70_Mode_Data".CRNT_MODE := 1; END_IF;
   "70_Mode_Data".AUT_RST_PLS.IN := "FirstScan";
END_REGION

REGION Network 2: Commanded Mode
   // Set mode as dictated by master PLC
   RUNG wire#powerrail
      Contact( "AlwaysTRUE" )
      I_Contact( "80_From_HMI".IGG_STND_ALN )
      Move(in := "50_CMND_DATA".CRNT_MODE, out1 => "70_Mode_Data".CRNT_MODE)
   END_RUNG
   // the same network as SCL:
   IF "AlwaysTRUE" AND NOT "80_From_HMI".IGG_STND_ALN THEN
       "70_Mode_Data".CRNT_MODE := "50_CMND_DATA".CRNT_MODE;
   END_IF;
END_REGION

REGION Network 3: Mode = Automatic
   // Automatic Mode
   RUNG wire#powerrail
      Contact( "80_From_HMI".IGG_STND_ALN )
      I_Contact( "80_From_HMI".FAT_Mode )
      Contact( "80_From_HMI".Request_Auto )
      wire#w1
      Move(in := 1, out1 => "70_Mode_Data".CRNT_MODE)
   END_RUNG
   RUNG wire#w1
      R_Coil( "120_FAT_FCS_DB".IN_FAT )
   END_RUNG
   // the same network as SCL:
   IF "80_From_HMI".IGG_STND_ALN AND NOT "80_From_HMI".FAT_Mode AND "80_From_HMI".Request_Auto THEN
       "70_Mode_Data".CRNT_MODE := 1;
       "120_FAT_FCS_DB".IN_FAT := FALSE;
   END_IF;
END_REGION

REGION Network 4: Mode = Manual
   // Manual Mode
   RUNG wire#powerrail
      Contact( "80_From_HMI".IGG_STND_ALN )
      I_Contact( "80_From_HMI".FAT_Mode )
      Contact( "80_From_HMI".Request_Manual )
      Move(in := 2, out1 => "70_Mode_Data".CRNT_MODE)
   END_RUNG
   // the same network as SCL:
   IF "80_From_HMI".IGG_STND_ALN AND NOT "80_From_HMI".FAT_Mode AND "80_From_HMI".Request_Manual THEN
       "70_Mode_Data".CRNT_MODE := 2;
   END_IF;
END_REGION

REGION Network 5: Mode = FAT Automatic
   // FAT Automatic Mode
   RUNG wire#powerrail
      Contact( "80_From_HMI".IGG_STND_ALN )
      Contact( "80_From_HMI".FAT_Mode )
      Contact( "80_From_HMI".Request_Auto )
      Move(in := 3, out1 => "70_Mode_Data".CRNT_MODE)
   END_RUNG
   // the same network as SCL:
   IF "80_From_HMI".IGG_STND_ALN AND "80_From_HMI".FAT_Mode AND "80_From_HMI".Request_Auto THEN
       "70_Mode_Data".CRNT_MODE := 3;
   END_IF;
END_REGION

REGION Network 6: Mode = FAT Manual
   // FAT Manual Mode
   RUNG wire#powerrail
      Contact( "80_From_HMI".IGG_STND_ALN )
      Contact( "80_From_HMI".FAT_Mode )
      Contact( "80_From_HMI".Request_Manual )
      Move(in := 4, out1 => "70_Mode_Data".CRNT_MODE)
   END_RUNG
   // the same network as SCL:
   IF "80_From_HMI".IGG_STND_ALN AND "80_From_HMI".FAT_Mode AND "80_From_HMI".Request_Manual THEN
       "70_Mode_Data".CRNT_MODE := 4;
   END_IF;
END_REGION
